DATA_BLOCK "DB149_KMI_FRA_Data"   // DB149
{ S7_Optimized_Access := 'FALSE' }
VERSION : 0.1
   VAR
      Signals_INT01 : Struct
         AP_ProgNr_Bit0 : Bool := FALSE;
         AP_ProgNr_Bit1 : Bool := FALSE;
         AP_ProgNr_Bit2 : Bool := FALSE;
         AP_ProgNr_Bit3 : Bool := FALSE;
         AP_ProgNr_Bit4 : Bool := FALSE;
         AP_ProgNr_Bit5 : Bool := FALSE;
         AP_ProgNr_Bit6 : Bool := FALSE;
         AP_ProgNr_Bit7 : Bool := FALSE;
         AP_OK : Bool := FALSE;
         AP_Strobe : Bool := FALSE;
         AP_Strobe_Inv : Bool := FALSE;
         AP_Shot : Bool := FALSE;
         AP_CP_forward : Bool := FALSE;
         AP_Filling : Bool := FALSE;
         AP_Res_0_6 : Bool := FALSE;
         AP_Res_0_7_1 : Bool := FALSE;
         PU_OK : Bool := FALSE;
         PU_Strobe_Quitt : Bool := FALSE;
         PU_Cycle_activ : Bool := FALSE;
         PU_Ready_for_shot : Bool := FALSE;
         PU_Shot_activ : Bool := FALSE;
         PU_Shot_End : Bool := FALSE;
         PU_Service_mode : Bool := TRUE;
         PU_CP_forward : Bool := FALSE;
         PU_Res_1_0 : Bool := FALSE;
         PU_Res_1_1 : Bool := FALSE;
         PU_Res_1_2 : Bool := FALSE;
         PU_Res_1_3 : Bool := FALSE;
         PU_Res_1_4 : Bool := FALSE;
         PU_Res_1_5 : Bool := FALSE;
         PU_Res_1_6 : Bool := FALSE;
         PU_Res_1_7 : Bool := FALSE;
         AP_Res_0_7 : Bool := FALSE;
      END_STRUCT;
      Measured_values_to_INT01 : Struct
         MH_Number : Byte := 16#01;
         Shot_Weight : Int := 16#1D40;
         Shot_Time : DInt := 16#0000_018D;
         Temperature_Poly : Int := 16#0794;
         Temperature_Iso : Int := 16#076C;
         Temperature_C3 : Int := 16#0000;
         Temperature_C4 : Int := 16#0000;
         Mix_Rate_Poly : Int := 16#2710;
         Mix_Rate_Iso : Int := 16#2F12;
         Mix_Rate_C3 : Int := 16#0000;
         Mix_Rate_C4 : Int := 16#0000;
         Pressure_Poly : Int := 16#466E;
         Pressure_Iso : Int := 16#44DE;
         Pressure_C3 : Int := 16#0000;
         Pressure_C4 : Int := 16#0000;
         Alarm_flow_K1 : Bool := FALSE;
         Alarm_flow_K2 : Bool := FALSE;
         Alarm_flow_K3 : Bool := FALSE;
         Alarm_flow_K4 : Bool := FALSE;
         Alarm_press_K1 : Bool := FALSE;
         Alarm_press_K2 : Bool := FALSE;
         Alarm_press_K3 : Bool := FALSE;
         Alarm_press_K4 : Bool := FALSE;
         Alarm_temp_K1 : Bool := FALSE;
         Alarm_temp_K2 : Bool := FALSE;
         Alarm_temp_K3 : Bool := FALSE;
         Alarm_temp_K4 : Bool := FALSE;
         Alarm_spare1 : Bool := FALSE;
         Alarm_spare2 : Bool := FALSE;
         Alarm_shottime : Bool := FALSE;
         Strobe_ProcessData : Bool := FALSE;
         Spare1 : Word := 16#0000;
         Spare2 : Word := 16#0000;
         Spare3 : Word := 16#0000;
         Spare4 : Word := 16#0000;
      END_STRUCT;
      Signals_INT02 : Struct
         AP_ProgNr_Bit0 : Bool := FALSE;
         AP_ProgNr_Bit1 : Bool := FALSE;
         AP_ProgNr_Bit2 : Bool := FALSE;
         AP_ProgNr_Bit3 : Bool := FALSE;
         AP_ProgNr_Bit4 : Bool := FALSE;
         AP_ProgNr_Bit5 : Bool := FALSE;
         AP_ProgNr_Bit6 : Bool := FALSE;
         AP_ProgNr_Bit7 : Bool := FALSE;
         AP_OK : Bool := FALSE;
         AP_Strobe : Bool := FALSE;
         AP_Strobe_Inv : Bool := FALSE;
         AP_Shot : Bool := FALSE;
         AP_CP_forward : Bool := FALSE;
         AP_Filling : Bool := FALSE;
         AP_Res_0_6 : Bool := FALSE;
         AP_Res_0_7_1 : Bool := FALSE;
         PU_OK : Bool := FALSE;
         PU_Strobe_Quitt : Bool := FALSE;
         PU_Cycle_activ : Bool := FALSE;
         PU_Ready_for_shot : Bool := FALSE;
         PU_Shot_activ : Bool := FALSE;
         PU_Shot_End : Bool := FALSE;
         PU_Service_mode : Bool := TRUE;
         PU_CP_forward : Bool := FALSE;
         PU_Res_1_0 : Bool := FALSE;
         PU_Res_1_1 : Bool := FALSE;
         PU_Res_1_2 : Bool := FALSE;
         PU_Res_1_3 : Bool := FALSE;
         PU_Res_1_4 : Bool := FALSE;
         PU_Res_1_5 : Bool := FALSE;
         PU_Res_1_6 : Bool := FALSE;
         PU_Res_1_7 : Bool := FALSE;
         AP_Res_0_7 : Bool := FALSE;
      END_STRUCT;
      Measured_values_to_INT02 : Struct
         MH_Number : Byte := 16#00;
         Shot_Weight : Int := 16#0000;
         Shot_Time : DInt := 16#0000_0000;
         Temperature_Poly : Int := 16#0000;
         Temperature_Iso : Int := 16#0000;
         Temperature_C3 : Int := 16#0000;
         Temperature_C4 : Int := 16#0000;
         Mix_Rate_Poly : Int := 16#0000;
         Mix_Rate_Iso : Int := 16#0000;
         Mix_Rate_C3 : Int := 16#0000;
         Mix_Rate_C4 : Int := 16#0000;
         Pressure_Poly : Int := 16#0000;
         Pressure_Iso : Int := 16#0000;
         Pressure_C3 : Int := 16#0000;
         Pressure_C4 : Int := 16#0000;
         Alarm_flow_K1 : Bool := FALSE;
         Alarm_flow_K2 : Bool := FALSE;
         Alarm_flow_K3 : Bool := FALSE;
         Alarm_flow_K4 : Bool := FALSE;
         Alarm_press_K1 : Bool := FALSE;
         Alarm_press_K2 : Bool := FALSE;
         Alarm_press_K3 : Bool := FALSE;
         Alarm_press_K4 : Bool := FALSE;
         Alarm_temp_K1 : Bool := FALSE;
         Alarm_temp_K2 : Bool := FALSE;
         Alarm_temp_K3 : Bool := FALSE;
         Alarm_temp_K4 : Bool := FALSE;
         Alarm_spare1 : Bool := FALSE;
         Alarm_spare2 : Bool := FALSE;
         Alarm_shottime : Bool := FALSE;
         Strobe_ProcessData : Bool := FALSE;
         Spare1 : Word := 16#0000;
         Spare2 : Word := 16#0000;
         Spare3 : Word := 16#0000;
         Spare4 : Word := 16#0000;
      END_STRUCT;
      Signals_INT03 : Struct
         AP_ProgNr_Bit0 : Bool := FALSE;
         AP_ProgNr_Bit1 : Bool := FALSE;
         AP_ProgNr_Bit2 : Bool := FALSE;
         AP_ProgNr_Bit3 : Bool := FALSE;
         AP_ProgNr_Bit4 : Bool := FALSE;
         AP_ProgNr_Bit5 : Bool := FALSE;
         AP_ProgNr_Bit6 : Bool := FALSE;
         AP_ProgNr_Bit7 : Bool := FALSE;
         AP_OK : Bool := FALSE;
         AP_Strobe : Bool := FALSE;
         AP_Strobe_Inv : Bool := FALSE;
         AP_Shot : Bool := FALSE;
         AP_CP_forward : Bool := FALSE;
         AP_Filling : Bool := FALSE;
         AP_Res_0_6 : Bool := FALSE;
         AP_Res_0_7_1 : Bool := FALSE;
         PU_OK : Bool := FALSE;
         PU_Strobe_Quitt : Bool := FALSE;
         PU_Cycle_activ : Bool := FALSE;
         PU_Ready_for_shot : Bool := FALSE;
         PU_Shot_activ : Bool := FALSE;
         PU_Shot_End : Bool := FALSE;
         PU_Service_mode : Bool := FALSE;
         PU_CP_forward : Bool := FALSE;
         PU_Res_1_0 : Bool := FALSE;
         PU_Res_1_1 : Bool := FALSE;
         PU_Res_1_2 : Bool := FALSE;
         PU_Res_1_3 : Bool := FALSE;
         PU_Res_1_4 : Bool := FALSE;
         PU_Res_1_5 : Bool := FALSE;
         PU_Res_1_6 : Bool := FALSE;
         PU_Res_1_7 : Bool := FALSE;
         AP_Res_0_7 : Bool := FALSE;
      END_STRUCT;
      Measured_values_to_INT03 : Struct
         MH_Number : Byte := 16#00;
         Shot_Weight : Int := 16#0000;
         Shot_Time : DInt := 16#0000_0000;
         Temperature_Poly : Int := 16#0000;
         Temperature_Iso : Int := 16#0000;
         Temperature_C3 : Int := 16#0000;
         Temperature_C4 : Int := 16#0000;
         Mix_Rate_Poly : Int := 16#0000;
         Mix_Rate_Iso : Int := 16#0000;
         Mix_Rate_C3 : Int := 16#0000;
         Mix_Rate_C4 : Int := 16#0000;
         Pressure_Poly : Int := 16#0000;
         Pressure_Iso : Int := 16#0000;
         Pressure_C3 : Int := 16#0000;
         Pressure_C4 : Int := 16#0000;
         Alarm_flow_K1 : Bool := FALSE;
         Alarm_flow_K2 : Bool := FALSE;
         Alarm_flow_K3 : Bool := FALSE;
         Alarm_flow_K4 : Bool := FALSE;
         Alarm_press_K1 : Bool := FALSE;
         Alarm_press_K2 : Bool := FALSE;
         Alarm_press_K3 : Bool := FALSE;
         Alarm_press_K4 : Bool := FALSE;
         Alarm_temp_K1 : Bool := FALSE;
         Alarm_temp_K2 : Bool := FALSE;
         Alarm_temp_K3 : Bool := FALSE;
         Alarm_temp_K4 : Bool := FALSE;
         Alarm_spare1 : Bool := FALSE;
         Alarm_spare2 : Bool := FALSE;
         Alarm_shottime : Bool := FALSE;
         Strobe_ProcessData : Bool := FALSE;
         Spare1 : Word := 16#0000;
         Spare2 : Word := 16#0000;
         Spare3 : Word := 16#0000;
         Spare4 : Word := 16#0000;
      END_STRUCT;
   END_VAR
BEGIN
END_DATA_BLOCK

DATA_BLOCK "DB_Zaehler_Anzeige"   // DB211
{ S7_Optimized_Access := 'FALSE' }
AUTHOR : AVP
NAME : MP270
VERSION : 0.1
   VAR
      ReadWriteDeviceNo : Int := 1;
      CopyDeviceNO : Int := 0;
      Read : Bool := FALSE;
      Write : Bool := FALSE;
      Copy : Bool := FALSE;
      Schichtwechsel : Bool := FALSE;
      ViewPreShift : Bool := FALSE;
      Gesamt : "Counter";
      "Counter" : Array[1..10] of "Counter";
      MH_Counter_ActualShift : Array[1..16] of Real;
      MH_Counter_PreShift : Array[1..16] of Real;
      MH_Counter_Reset : Array[1..16] of Real;
      MH_Counter_NonReset : Array[1..16] of Real;
   END_VAR
BEGIN
   Gesamt.Anzahl := 0;
   Gesamt.Verbrauch_K1 := 0.0;
   Gesamt.Verbrauch_K2 := 0.0;
   Gesamt.Verbrauch_K3 := 0.0;
   Gesamt.Verbrauch_K4 := 0.0;
   Gesamt.Verbrauch_K5 := 0.0;
   Gesamt.Verbrauch_K6 := 0.0;
   Gesamt.Verbrauch_K7 := 0.0;
   Gesamt.Verbrauch_K8 := 0.0;
   "Counter"[1].Anzahl := 0;
   "Counter"[1].Verbrauch_K1 := 0.0;
   "Counter"[1].Verbrauch_K2 := 0.0;
   "Counter"[1].Verbrauch_K3 := 0.0;
   "Counter"[1].Verbrauch_K4 := 0.0;
   "Counter"[1].Verbrauch_K5 := 0.0;
   "Counter"[1].Verbrauch_K6 := 0.0;
   "Counter"[1].Verbrauch_K7 := 0.0;
   "Counter"[1].Verbrauch_K8 := 0.0;
   "Counter"[2].Anzahl := 0;
   "Counter"[2].Verbrauch_K1 := 0.0;
   "Counter"[2].Verbrauch_K2 := 0.0;
   "Counter"[2].Verbrauch_K3 := 0.0;
   "Counter"[2].Verbrauch_K4 := 0.0;
   "Counter"[2].Verbrauch_K5 := 0.0;
   "Counter"[2].Verbrauch_K6 := 0.0;
   "Counter"[2].Verbrauch_K7 := 0.0;
   "Counter"[2].Verbrauch_K8 := 0.0;
   "Counter"[3].Anzahl := 0;
   "Counter"[3].Verbrauch_K1 := 0.0;
   "Counter"[3].Verbrauch_K2 := 0.0;
   "Counter"[3].Verbrauch_K3 := 0.0;
   "Counter"[3].Verbrauch_K4 := 0.0;
   "Counter"[3].Verbrauch_K5 := 0.0;
   "Counter"[3].Verbrauch_K6 := 0.0;
   "Counter"[3].Verbrauch_K7 := 0.0;
   "Counter"[3].Verbrauch_K8 := 0.0;
   "Counter"[4].Anzahl := 0;
   "Counter"[4].Verbrauch_K1 := 0.0;
   "Counter"[4].Verbrauch_K2 := 0.0;
   "Counter"[4].Verbrauch_K3 := 0.0;
   "Counter"[4].Verbrauch_K4 := 0.0;
   "Counter"[4].Verbrauch_K5 := 0.0;
   "Counter"[4].Verbrauch_K6 := 0.0;
   "Counter"[4].Verbrauch_K7 := 0.0;
   "Counter"[4].Verbrauch_K8 := 0.0;
   "Counter"[5].Anzahl := 0;
   "Counter"[5].Verbrauch_K1 := 0.0;
   "Counter"[5].Verbrauch_K2 := 0.0;
   "Counter"[5].Verbrauch_K3 := 0.0;
   "Counter"[5].Verbrauch_K4 := 0.0;
   "Counter"[5].Verbrauch_K5 := 0.0;
   "Counter"[5].Verbrauch_K6 := 0.0;
   "Counter"[5].Verbrauch_K7 := 0.0;
   "Counter"[5].Verbrauch_K8 := 0.0;
   "Counter"[6].Anzahl := 0;
   "Counter"[6].Verbrauch_K1 := 0.0;
   "Counter"[6].Verbrauch_K2 := 0.0;
   "Counter"[6].Verbrauch_K3 := 0.0;
   "Counter"[6].Verbrauch_K4 := 0.0;
   "Counter"[6].Verbrauch_K5 := 0.0;
   "Counter"[6].Verbrauch_K6 := 0.0;
   "Counter"[6].Verbrauch_K7 := 0.0;
   "Counter"[6].Verbrauch_K8 := 0.0;
   "Counter"[7].Anzahl := 0;
   "Counter"[7].Verbrauch_K1 := 0.0;
   "Counter"[7].Verbrauch_K2 := 0.0;
   "Counter"[7].Verbrauch_K3 := 0.0;
   "Counter"[7].Verbrauch_K4 := 0.0;
   "Counter"[7].Verbrauch_K5 := 0.0;
   "Counter"[7].Verbrauch_K6 := 0.0;
   "Counter"[7].Verbrauch_K7 := 0.0;
   "Counter"[7].Verbrauch_K8 := 0.0;
   "Counter"[8].Anzahl := 0;
   "Counter"[8].Verbrauch_K1 := 0.0;
   "Counter"[8].Verbrauch_K2 := 0.0;
   "Counter"[8].Verbrauch_K3 := 0.0;
   "Counter"[8].Verbrauch_K4 := 0.0;
   "Counter"[8].Verbrauch_K5 := 0.0;
   "Counter"[8].Verbrauch_K6 := 0.0;
   "Counter"[8].Verbrauch_K7 := 0.0;
   "Counter"[8].Verbrauch_K8 := 0.0;
   "Counter"[9].Anzahl := 0;
   "Counter"[9].Verbrauch_K1 := 0.0;
   "Counter"[9].Verbrauch_K2 := 0.0;
   "Counter"[9].Verbrauch_K3 := 0.0;
   "Counter"[9].Verbrauch_K4 := 0.0;
   "Counter"[9].Verbrauch_K5 := 0.0;
   "Counter"[9].Verbrauch_K6 := 0.0;
   "Counter"[9].Verbrauch_K7 := 0.0;
   "Counter"[9].Verbrauch_K8 := 0.0;
   "Counter"[10].Anzahl := 0;
   "Counter"[10].Verbrauch_K1 := 0.0;
   "Counter"[10].Verbrauch_K2 := 0.0;
   "Counter"[10].Verbrauch_K3 := 0.0;
   "Counter"[10].Verbrauch_K4 := 0.0;
   "Counter"[10].Verbrauch_K5 := 0.0;
   "Counter"[10].Verbrauch_K6 := 0.0;
   "Counter"[10].Verbrauch_K7 := 0.0;
   "Counter"[10].Verbrauch_K8 := 0.0;
   MH_Counter_ActualShift[1] := 0.0;
   MH_Counter_ActualShift[2] := 0.0;
   MH_Counter_ActualShift[3] := 0.0;
   MH_Counter_ActualShift[4] := 0.0;
   MH_Counter_ActualShift[5] := 0.0;
   MH_Counter_ActualShift[6] := 0.0;
   MH_Counter_ActualShift[7] := 0.0;
   MH_Counter_ActualShift[8] := 0.0;
   MH_Counter_ActualShift[9] := 0.0;
   MH_Counter_ActualShift[10] := 0.0;
   MH_Counter_ActualShift[11] := 0.0;
   MH_Counter_ActualShift[12] := 0.0;
   MH_Counter_ActualShift[13] := 0.0;
   MH_Counter_ActualShift[14] := 0.0;
   MH_Counter_ActualShift[15] := 0.0;
   MH_Counter_ActualShift[16] := 0.0;
   MH_Counter_PreShift[1] := 0.0;
   MH_Counter_PreShift[2] := 0.0;
   MH_Counter_PreShift[3] := 0.0;
   MH_Counter_PreShift[4] := 0.0;
   MH_Counter_PreShift[5] := 0.0;
   MH_Counter_PreShift[6] := 0.0;
   MH_Counter_PreShift[7] := 0.0;
   MH_Counter_PreShift[8] := 0.0;
   MH_Counter_PreShift[9] := 0.0;
   MH_Counter_PreShift[10] := 0.0;
   MH_Counter_PreShift[11] := 0.0;
   MH_Counter_PreShift[12] := 0.0;
   MH_Counter_PreShift[13] := 0.0;
   MH_Counter_PreShift[14] := 0.0;
   MH_Counter_PreShift[15] := 0.0;
   MH_Counter_PreShift[16] := 0.0;
   MH_Counter_Reset[1] := 0.0;
   MH_Counter_Reset[2] := 0.0;
   MH_Counter_Reset[3] := 0.0;
   MH_Counter_Reset[4] := 0.0;
   MH_Counter_Reset[5] := 0.0;
   MH_Counter_Reset[6] := 0.0;
   MH_Counter_Reset[7] := 0.0;
   MH_Counter_Reset[8] := 0.0;
   MH_Counter_Reset[9] := 0.0;
   MH_Counter_Reset[10] := 0.0;
   MH_Counter_Reset[11] := 0.0;
   MH_Counter_Reset[12] := 0.0;
   MH_Counter_Reset[13] := 0.0;
   MH_Counter_Reset[14] := 0.0;
   MH_Counter_Reset[15] := 0.0;
   MH_Counter_Reset[16] := 0.0;
   MH_Counter_NonReset[1] := 0.0;
   MH_Counter_NonReset[2] := 0.0;
   MH_Counter_NonReset[3] := 0.0;
   MH_Counter_NonReset[4] := 0.0;
   MH_Counter_NonReset[5] := 0.0;
   MH_Counter_NonReset[6] := 0.0;
   MH_Counter_NonReset[7] := 0.0;
   MH_Counter_NonReset[8] := 0.0;
   MH_Counter_NonReset[9] := 0.0;
   MH_Counter_NonReset[10] := 0.0;
   MH_Counter_NonReset[11] := 0.0;
   MH_Counter_NonReset[12] := 0.0;
   MH_Counter_NonReset[13] := 0.0;
   MH_Counter_NonReset[14] := 0.0;
   MH_Counter_NonReset[15] := 0.0;
   MH_Counter_NonReset[16] := 0.0;
END_DATA_BLOCK

DATA_BLOCK "DB_Zaehler_Schicht_aktuell"   // DB212
{ S7_Optimized_Access := 'FALSE' }
AUTHOR : AVP
NAME : MP270
VERSION : 0.1
   VAR
      Gesamt : "Counter";
      "Counter" : Array[1..120] of "Counter";
      MH_Counter : Array[1..16] of Real;
   END_VAR
BEGIN
   Gesamt.Anzahl := 0;
   Gesamt.Verbrauch_K1 := 0.0;
   Gesamt.Verbrauch_K2 := 0.0;
   Gesamt.Verbrauch_K3 := 0.0;
   Gesamt.Verbrauch_K4 := 0.0;
   Gesamt.Verbrauch_K5 := 0.0;
   Gesamt.Verbrauch_K6 := 0.0;
   Gesamt.Verbrauch_K7 := 0.0;
   Gesamt.Verbrauch_K8 := 0.0;
   "Counter"[1].Anzahl := 0;
   "Counter"[1].Verbrauch_K1 := 0.0;
   "Counter"[1].Verbrauch_K2 := 0.0;
   "Counter"[1].Verbrauch_K3 := 0.0;
   "Counter"[1].Verbrauch_K4 := 0.0;
   "Counter"[1].Verbrauch_K5 := 0.0;
   "Counter"[1].Verbrauch_K6 := 0.0;
   "Counter"[1].Verbrauch_K7 := 0.0;
   "Counter"[1].Verbrauch_K8 := 0.0;
   "Counter"[2].Anzahl := 0;
   "Counter"[2].Verbrauch_K1 := 0.0;
   "Counter"[2].Verbrauch_K2 := 0.0;
   "Counter"[2].Verbrauch_K3 := 0.0;
   "Counter"[2].Verbrauch_K4 := 0.0;
   "Counter"[2].Verbrauch_K5 := 0.0;
   "Counter"[2].Verbrauch_K6 := 0.0;
   "Counter"[2].Verbrauch_K7 := 0.0;
   "Counter"[2].Verbrauch_K8 := 0.0;
   "Counter"[3].Anzahl := 0;
   "Counter"[3].Verbrauch_K1 := 0.0;
   "Counter"[3].Verbrauch_K2 := 0.0;
   "Counter"[3].Verbrauch_K3 := 0.0;
   "Counter"[3].Verbrauch_K4 := 0.0;
   "Counter"[3].Verbrauch_K5 := 0.0;
   "Counter"[3].Verbrauch_K6 := 0.0;
   "Counter"[3].Verbrauch_K7 := 0.0;
   "Counter"[3].Verbrauch_K8 := 0.0;
   "Counter"[4].Anzahl := 0;
   "Counter"[4].Verbrauch_K1 := 0.0;
   "Counter"[4].Verbrauch_K2 := 0.0;
   "Counter"[4].Verbrauch_K3 := 0.0;
   "Counter"[4].Verbrauch_K4 := 0.0;
   "Counter"[4].Verbrauch_K5 := 0.0;
   "Counter"[4].Verbrauch_K6 := 0.0;
   "Counter"[4].Verbrauch_K7 := 0.0;
   "Counter"[4].Verbrauch_K8 := 0.0;
   "Counter"[5].Anzahl := 0;
   "Counter"[5].Verbrauch_K1 := 0.0;
   "Counter"[5].Verbrauch_K2 := 0.0;
   "Counter"[5].Verbrauch_K3 := 0.0;
   "Counter"[5].Verbrauch_K4 := 0.0;
   "Counter"[5].Verbrauch_K5 := 0.0;
   "Counter"[5].Verbrauch_K6 := 0.0;
   "Counter"[5].Verbrauch_K7 := 0.0;
   "Counter"[5].Verbrauch_K8 := 0.0;
   "Counter"[6].Anzahl := 0;
   "Counter"[6].Verbrauch_K1 := 0.0;
   "Counter"[6].Verbrauch_K2 := 0.0;
   "Counter"[6].Verbrauch_K3 := 0.0;
   "Counter"[6].Verbrauch_K4 := 0.0;
   "Counter"[6].Verbrauch_K5 := 0.0;
   "Counter"[6].Verbrauch_K6 := 0.0;
   "Counter"[6].Verbrauch_K7 := 0.0;
   "Counter"[6].Verbrauch_K8 := 0.0;
   "Counter"[7].Anzahl := 0;
   "Counter"[7].Verbrauch_K1 := 0.0;
   "Counter"[7].Verbrauch_K2 := 0.0;
   "Counter"[7].Verbrauch_K3 := 0.0;
   "Counter"[7].Verbrauch_K4 := 0.0;
   "Counter"[7].Verbrauch_K5 := 0.0;
   "Counter"[7].Verbrauch_K6 := 0.0;
   "Counter"[7].Verbrauch_K7 := 0.0;
   "Counter"[7].Verbrauch_K8 := 0.0;
   "Counter"[8].Anzahl := 0;
   "Counter"[8].Verbrauch_K1 := 0.0;
   "Counter"[8].Verbrauch_K2 := 0.0;
   "Counter"[8].Verbrauch_K3 := 0.0;
   "Counter"[8].Verbrauch_K4 := 0.0;
   "Counter"[8].Verbrauch_K5 := 0.0;
   "Counter"[8].Verbrauch_K6 := 0.0;
   "Counter"[8].Verbrauch_K7 := 0.0;
   "Counter"[8].Verbrauch_K8 := 0.0;
   "Counter"[9].Anzahl := 0;
   "Counter"[9].Verbrauch_K1 := 0.0;
   "Counter"[9].Verbrauch_K2 := 0.0;
   "Counter"[9].Verbrauch_K3 := 0.0;
   "Counter"[9].Verbrauch_K4 := 0.0;
   "Counter"[9].Verbrauch_K5 := 0.0;
   "Counter"[9].Verbrauch_K6 := 0.0;
   "Counter"[9].Verbrauch_K7 := 0.0;
   "Counter"[9].Verbrauch_K8 := 0.0;
   "Counter"[10].Anzahl := 0;
   "Counter"[10].Verbrauch_K1 := 0.0;
   "Counter"[10].Verbrauch_K2 := 0.0;
   "Counter"[10].Verbrauch_K3 := 0.0;
   "Counter"[10].Verbrauch_K4 := 0.0;
   "Counter"[10].Verbrauch_K5 := 0.0;
   "Counter"[10].Verbrauch_K6 := 0.0;
   "Counter"[10].Verbrauch_K7 := 0.0;
   "Counter"[10].Verbrauch_K8 := 0.0;
   "Counter"[11].Anzahl := 0;
   "Counter"[11].Verbrauch_K1 := 0.0;
   "Counter"[11].Verbrauch_K2 := 0.0;
   "Counter"[11].Verbrauch_K3 := 0.0;
   "Counter"[11].Verbrauch_K4 := 0.0;
   "Counter"[11].Verbrauch_K5 := 0.0;
   "Counter"[11].Verbrauch_K6 := 0.0;
   "Counter"[11].Verbrauch_K7 := 0.0;
   "Counter"[11].Verbrauch_K8 := 0.0;
   "Counter"[12].Anzahl := 0;
   "Counter"[12].Verbrauch_K1 := 0.0;
   "Counter"[12].Verbrauch_K2 := 0.0;
   "Counter"[12].Verbrauch_K3 := 0.0;
   "Counter"[12].Verbrauch_K4 := 0.0;
   "Counter"[12].Verbrauch_K5 := 0.0;
   "Counter"[12].Verbrauch_K6 := 0.0;
   "Counter"[12].Verbrauch_K7 := 0.0;
   "Counter"[12].Verbrauch_K8 := 0.0;
   "Counter"[13].Anzahl := 0;
   "Counter"[13].Verbrauch_K1 := 0.0;
   "Counter"[13].Verbrauch_K2 := 0.0;
   "Counter"[13].Verbrauch_K3 := 0.0;
   "Counter"[13].Verbrauch_K4 := 0.0;
   "Counter"[13].Verbrauch_K5 := 0.0;
   "Counter"[13].Verbrauch_K6 := 0.0;
   "Counter"[13].Verbrauch_K7 := 0.0;
   "Counter"[13].Verbrauch_K8 := 0.0;
   "Counter"[14].Anzahl := 0;
   "Counter"[14].Verbrauch_K1 := 0.0;
   "Counter"[14].Verbrauch_K2 := 0.0;
   "Counter"[14].Verbrauch_K3 := 0.0;
   "Counter"[14].Verbrauch_K4 := 0.0;
   "Counter"[14].Verbrauch_K5 := 0.0;
   "Counter"[14].Verbrauch_K6 := 0.0;
   "Counter"[14].Verbrauch_K7 := 0.0;
   "Counter"[14].Verbrauch_K8 := 0.0;
   "Counter"[15].Anzahl := 0;
   "Counter"[15].Verbrauch_K1 := 0.0;
   "Counter"[15].Verbrauch_K2 := 0.0;
   "Counter"[15].Verbrauch_K3 := 0.0;
   "Counter"[15].Verbrauch_K4 := 0.0;
   "Counter"[15].Verbrauch_K5 := 0.0;
   "Counter"[15].Verbrauch_K6 := 0.0;
   "Counter"[15].Verbrauch_K7 := 0.0;
   "Counter"[15].Verbrauch_K8 := 0.0;
   "Counter"[16].Anzahl := 0;
   "Counter"[16].Verbrauch_K1 := 0.0;
   "Counter"[16].Verbrauch_K2 := 0.0;
   "Counter"[16].Verbrauch_K3 := 0.0;
   "Counter"[16].Verbrauch_K4 := 0.0;
   "Counter"[16].Verbrauch_K5 := 0.0;
   "Counter"[16].Verbrauch_K6 := 0.0;
   "Counter"[16].Verbrauch_K7 := 0.0;
   "Counter"[16].Verbrauch_K8 := 0.0;
   "Counter"[17].Anzahl := 0;
   "Counter"[17].Verbrauch_K1 := 0.0;
   "Counter"[17].Verbrauch_K2 := 0.0;
   "Counter"[17].Verbrauch_K3 := 0.0;
   "Counter"[17].Verbrauch_K4 := 0.0;
   "Counter"[17].Verbrauch_K5 := 0.0;
   "Counter"[17].Verbrauch_K6 := 0.0;
   "Counter"[17].Verbrauch_K7 := 0.0;
   "Counter"[17].Verbrauch_K8 := 0.0;
   "Counter"[18].Anzahl := 0;
   "Counter"[18].Verbrauch_K1 := 0.0;
   "Counter"[18].Verbrauch_K2 := 0.0;
   "Counter"[18].Verbrauch_K3 := 0.0;
   "Counter"[18].Verbrauch_K4 := 0.0;
   "Counter"[18].Verbrauch_K5 := 0.0;
   "Counter"[18].Verbrauch_K6 := 0.0;
   "Counter"[18].Verbrauch_K7 := 0.0;
   "Counter"[18].Verbrauch_K8 := 0.0;
   "Counter"[19].Anzahl := 0;
   "Counter"[19].Verbrauch_K1 := 0.0;
   "Counter"[19].Verbrauch_K2 := 0.0;
   "Counter"[19].Verbrauch_K3 := 0.0;
   "Counter"[19].Verbrauch_K4 := 0.0;
   "Counter"[19].Verbrauch_K5 := 0.0;
   "Counter"[19].Verbrauch_K6 := 0.0;
   "Counter"[19].Verbrauch_K7 := 0.0;
   "Counter"[19].Verbrauch_K8 := 0.0;
   "Counter"[20].Anzahl := 0;
   "Counter"[20].Verbrauch_K1 := 0.0;
   "Counter"[20].Verbrauch_K2 := 0.0;
   "Counter"[20].Verbrauch_K3 := 0.0;
   "Counter"[20].Verbrauch_K4 := 0.0;
   "Counter"[20].Verbrauch_K5 := 0.0;
   "Counter"[20].Verbrauch_K6 := 0.0;
   "Counter"[20].Verbrauch_K7 := 0.0;
   "Counter"[20].Verbrauch_K8 := 0.0;
   "Counter"[21].Anzahl := 0;
   "Counter"[21].Verbrauch_K1 := 0.0;
   "Counter"[21].Verbrauch_K2 := 0.0;
   "Counter"[21].Verbrauch_K3 := 0.0;
   "Counter"[21].Verbrauch_K4 := 0.0;
   "Counter"[21].Verbrauch_K5 := 0.0;
   "Counter"[21].Verbrauch_K6 := 0.0;
   "Counter"[21].Verbrauch_K7 := 0.0;
   "Counter"[21].Verbrauch_K8 := 0.0;
   "Counter"[22].Anzahl := 0;
   "Counter"[22].Verbrauch_K1 := 0.0;
   // 905 more start values not shown
END_DATA_BLOCK

DATA_BLOCK "DB_Zaehler_Schicht_Vorherige"   // DB213
{ S7_Optimized_Access := 'FALSE' }
VERSION : 0.1
   VAR
      Gesamt : "Counter";
      "Counter" : Array[1..120] of "Counter";
      MH_Counter : Array[1..16] of Real;
   END_VAR
BEGIN
   Gesamt.Anzahl := 0;
   Gesamt.Verbrauch_K1 := 0.0;
   Gesamt.Verbrauch_K2 := 0.0;
   Gesamt.Verbrauch_K3 := 0.0;
   Gesamt.Verbrauch_K4 := 0.0;
   Gesamt.Verbrauch_K5 := 0.0;
   Gesamt.Verbrauch_K6 := 0.0;
   Gesamt.Verbrauch_K7 := 0.0;
   Gesamt.Verbrauch_K8 := 0.0;
   "Counter"[1].Anzahl := 0;
   "Counter"[1].Verbrauch_K1 := 0.0;
   "Counter"[1].Verbrauch_K2 := 0.0;
   "Counter"[1].Verbrauch_K3 := 0.0;
   "Counter"[1].Verbrauch_K4 := 0.0;
   "Counter"[1].Verbrauch_K5 := 0.0;
   "Counter"[1].Verbrauch_K6 := 0.0;
   "Counter"[1].Verbrauch_K7 := 0.0;
   "Counter"[1].Verbrauch_K8 := 0.0;
   "Counter"[2].Anzahl := 0;
   "Counter"[2].Verbrauch_K1 := 0.0;
   "Counter"[2].Verbrauch_K2 := 0.0;
   "Counter"[2].Verbrauch_K3 := 0.0;
   "Counter"[2].Verbrauch_K4 := 0.0;
   "Counter"[2].Verbrauch_K5 := 0.0;
   "Counter"[2].Verbrauch_K6 := 0.0;
   "Counter"[2].Verbrauch_K7 := 0.0;
   "Counter"[2].Verbrauch_K8 := 0.0;
   "Counter"[3].Anzahl := 0;
   "Counter"[3].Verbrauch_K1 := 0.0;
   "Counter"[3].Verbrauch_K2 := 0.0;
   "Counter"[3].Verbrauch_K3 := 0.0;
   "Counter"[3].Verbrauch_K4 := 0.0;
   "Counter"[3].Verbrauch_K5 := 0.0;
   "Counter"[3].Verbrauch_K6 := 0.0;
   "Counter"[3].Verbrauch_K7 := 0.0;
   "Counter"[3].Verbrauch_K8 := 0.0;
   "Counter"[4].Anzahl := 0;
   "Counter"[4].Verbrauch_K1 := 0.0;
   "Counter"[4].Verbrauch_K2 := 0.0;
   "Counter"[4].Verbrauch_K3 := 0.0;
   "Counter"[4].Verbrauch_K4 := 0.0;
   "Counter"[4].Verbrauch_K5 := 0.0;
   "Counter"[4].Verbrauch_K6 := 0.0;
   "Counter"[4].Verbrauch_K7 := 0.0;
   "Counter"[4].Verbrauch_K8 := 0.0;
   "Counter"[5].Anzahl := 0;
   "Counter"[5].Verbrauch_K1 := 0.0;
   "Counter"[5].Verbrauch_K2 := 0.0;
   "Counter"[5].Verbrauch_K3 := 0.0;
   "Counter"[5].Verbrauch_K4 := 0.0;
   "Counter"[5].Verbrauch_K5 := 0.0;
   "Counter"[5].Verbrauch_K6 := 0.0;
   "Counter"[5].Verbrauch_K7 := 0.0;
   "Counter"[5].Verbrauch_K8 := 0.0;
   "Counter"[6].Anzahl := 0;
   "Counter"[6].Verbrauch_K1 := 0.0;
   "Counter"[6].Verbrauch_K2 := 0.0;
   "Counter"[6].Verbrauch_K3 := 0.0;
   "Counter"[6].Verbrauch_K4 := 0.0;
   "Counter"[6].Verbrauch_K5 := 0.0;
   "Counter"[6].Verbrauch_K6 := 0.0;
   "Counter"[6].Verbrauch_K7 := 0.0;
   "Counter"[6].Verbrauch_K8 := 0.0;
   "Counter"[7].Anzahl := 0;
   "Counter"[7].Verbrauch_K1 := 0.0;
   "Counter"[7].Verbrauch_K2 := 0.0;
   "Counter"[7].Verbrauch_K3 := 0.0;
   "Counter"[7].Verbrauch_K4 := 0.0;
   "Counter"[7].Verbrauch_K5 := 0.0;
   "Counter"[7].Verbrauch_K6 := 0.0;
   "Counter"[7].Verbrauch_K7 := 0.0;
   "Counter"[7].Verbrauch_K8 := 0.0;
   "Counter"[8].Anzahl := 0;
   "Counter"[8].Verbrauch_K1 := 0.0;
   "Counter"[8].Verbrauch_K2 := 0.0;
   "Counter"[8].Verbrauch_K3 := 0.0;
   "Counter"[8].Verbrauch_K4 := 0.0;
   "Counter"[8].Verbrauch_K5 := 0.0;
   "Counter"[8].Verbrauch_K6 := 0.0;
   "Counter"[8].Verbrauch_K7 := 0.0;
   "Counter"[8].Verbrauch_K8 := 0.0;
   "Counter"[9].Anzahl := 0;
   "Counter"[9].Verbrauch_K1 := 0.0;
   "Counter"[9].Verbrauch_K2 := 0.0;
   "Counter"[9].Verbrauch_K3 := 0.0;
   "Counter"[9].Verbrauch_K4 := 0.0;
   "Counter"[9].Verbrauch_K5 := 0.0;
   "Counter"[9].Verbrauch_K6 := 0.0;
   "Counter"[9].Verbrauch_K7 := 0.0;
   "Counter"[9].Verbrauch_K8 := 0.0;
   "Counter"[10].Anzahl := 0;
   "Counter"[10].Verbrauch_K1 := 0.0;
   "Counter"[10].Verbrauch_K2 := 0.0;
   "Counter"[10].Verbrauch_K3 := 0.0;
   "Counter"[10].Verbrauch_K4 := 0.0;
   "Counter"[10].Verbrauch_K5 := 0.0;
   "Counter"[10].Verbrauch_K6 := 0.0;
   "Counter"[10].Verbrauch_K7 := 0.0;
   "Counter"[10].Verbrauch_K8 := 0.0;
   "Counter"[11].Anzahl := 0;
   "Counter"[11].Verbrauch_K1 := 0.0;
   "Counter"[11].Verbrauch_K2 := 0.0;
   "Counter"[11].Verbrauch_K3 := 0.0;
   "Counter"[11].Verbrauch_K4 := 0.0;
   "Counter"[11].Verbrauch_K5 := 0.0;
   "Counter"[11].Verbrauch_K6 := 0.0;
   "Counter"[11].Verbrauch_K7 := 0.0;
   "Counter"[11].Verbrauch_K8 := 0.0;
   "Counter"[12].Anzahl := 0;
   "Counter"[12].Verbrauch_K1 := 0.0;
   "Counter"[12].Verbrauch_K2 := 0.0;
   "Counter"[12].Verbrauch_K3 := 0.0;
   "Counter"[12].Verbrauch_K4 := 0.0;
   "Counter"[12].Verbrauch_K5 := 0.0;
   "Counter"[12].Verbrauch_K6 := 0.0;
   "Counter"[12].Verbrauch_K7 := 0.0;
   "Counter"[12].Verbrauch_K8 := 0.0;
   "Counter"[13].Anzahl := 0;
   "Counter"[13].Verbrauch_K1 := 0.0;
   "Counter"[13].Verbrauch_K2 := 0.0;
   "Counter"[13].Verbrauch_K3 := 0.0;
   "Counter"[13].Verbrauch_K4 := 0.0;
   "Counter"[13].Verbrauch_K5 := 0.0;
   "Counter"[13].Verbrauch_K6 := 0.0;
   "Counter"[13].Verbrauch_K7 := 0.0;
   "Counter"[13].Verbrauch_K8 := 0.0;
   "Counter"[14].Anzahl := 0;
   "Counter"[14].Verbrauch_K1 := 0.0;
   "Counter"[14].Verbrauch_K2 := 0.0;
   "Counter"[14].Verbrauch_K3 := 0.0;
   "Counter"[14].Verbrauch_K4 := 0.0;
   "Counter"[14].Verbrauch_K5 := 0.0;
   "Counter"[14].Verbrauch_K6 := 0.0;
   "Counter"[14].Verbrauch_K7 := 0.0;
   "Counter"[14].Verbrauch_K8 := 0.0;
   "Counter"[15].Anzahl := 0;
   "Counter"[15].Verbrauch_K1 := 0.0;
   "Counter"[15].Verbrauch_K2 := 0.0;
   "Counter"[15].Verbrauch_K3 := 0.0;
   "Counter"[15].Verbrauch_K4 := 0.0;
   "Counter"[15].Verbrauch_K5 := 0.0;
   "Counter"[15].Verbrauch_K6 := 0.0;
   "Counter"[15].Verbrauch_K7 := 0.0;
   "Counter"[15].Verbrauch_K8 := 0.0;
   "Counter"[16].Anzahl := 0;
   "Counter"[16].Verbrauch_K1 := 0.0;
   "Counter"[16].Verbrauch_K2 := 0.0;
   "Counter"[16].Verbrauch_K3 := 0.0;
   "Counter"[16].Verbrauch_K4 := 0.0;
   "Counter"[16].Verbrauch_K5 := 0.0;
   "Counter"[16].Verbrauch_K6 := 0.0;
   "Counter"[16].Verbrauch_K7 := 0.0;
   "Counter"[16].Verbrauch_K8 := 0.0;
   "Counter"[17].Anzahl := 0;
   "Counter"[17].Verbrauch_K1 := 0.0;
   "Counter"[17].Verbrauch_K2 := 0.0;
   "Counter"[17].Verbrauch_K3 := 0.0;
   "Counter"[17].Verbrauch_K4 := 0.0;
   "Counter"[17].Verbrauch_K5 := 0.0;
   "Counter"[17].Verbrauch_K6 := 0.0;
   "Counter"[17].Verbrauch_K7 := 0.0;
   "Counter"[17].Verbrauch_K8 := 0.0;
   "Counter"[18].Anzahl := 0;
   "Counter"[18].Verbrauch_K1 := 0.0;
   "Counter"[18].Verbrauch_K2 := 0.0;
   "Counter"[18].Verbrauch_K3 := 0.0;
   "Counter"[18].Verbrauch_K4 := 0.0;
   "Counter"[18].Verbrauch_K5 := 0.0;
   "Counter"[18].Verbrauch_K6 := 0.0;
   "Counter"[18].Verbrauch_K7 := 0.0;
   "Counter"[18].Verbrauch_K8 := 0.0;
   "Counter"[19].Anzahl := 0;
   "Counter"[19].Verbrauch_K1 := 0.0;
   "Counter"[19].Verbrauch_K2 := 0.0;
   "Counter"[19].Verbrauch_K3 := 0.0;
   "Counter"[19].Verbrauch_K4 := 0.0;
   "Counter"[19].Verbrauch_K5 := 0.0;
   "Counter"[19].Verbrauch_K6 := 0.0;
   "Counter"[19].Verbrauch_K7 := 0.0;
   "Counter"[19].Verbrauch_K8 := 0.0;
   "Counter"[20].Anzahl := 0;
   "Counter"[20].Verbrauch_K1 := 0.0;
   "Counter"[20].Verbrauch_K2 := 0.0;
   "Counter"[20].Verbrauch_K3 := 0.0;
   "Counter"[20].Verbrauch_K4 := 0.0;
   "Counter"[20].Verbrauch_K5 := 0.0;
   "Counter"[20].Verbrauch_K6 := 0.0;
   "Counter"[20].Verbrauch_K7 := 0.0;
   "Counter"[20].Verbrauch_K8 := 0.0;
   "Counter"[21].Anzahl := 0;
   "Counter"[21].Verbrauch_K1 := 0.0;
   "Counter"[21].Verbrauch_K2 := 0.0;
   "Counter"[21].Verbrauch_K3 := 0.0;
   "Counter"[21].Verbrauch_K4 := 0.0;
   "Counter"[21].Verbrauch_K5 := 0.0;
   "Counter"[21].Verbrauch_K6 := 0.0;
   "Counter"[21].Verbrauch_K7 := 0.0;
   "Counter"[21].Verbrauch_K8 := 0.0;
   "Counter"[22].Anzahl := 0;
   "Counter"[22].Verbrauch_K1 := 0.0;
   // 905 more start values not shown
END_DATA_BLOCK

DATA_BLOCK "DB315_ShotadjustS"   // DB315
TITLE = Shot time correction for each partshot of a tool
{ S7_Optimized_Access := 'FALSE' }
VERSION : 0.1
   VAR
      Tool : Array[0..120] of "UDT315_ShotadjustS";   // Shot time correction for each partshot of a tool
   END_VAR
BEGIN
   Tool[0].PS1 := 0.0;
END_DATA_BLOCK

DATA_BLOCK "DB601_PV_Plunger"   // DB601
TITLE = Process values of metering plunger
{ S7_Optimized_Access := 'FALSE' }
AUTHOR : KT242
VERSION : 0.1
   VAR
      ReadWriteDeviceNo : Int;
      CopyDeviceNO : Int;
      Read : Bool;
      Write : Bool;
      Copy : Bool;
      Component : Array[0..12] of "UDT509_PV_Plunger";
   END_VAR
BEGIN
END_DATA_BLOCK

DATA_BLOCK "DB602_PV_Tank"   // DB602
TITLE = Process values of tanks
{ S7_Optimized_Access := 'FALSE' }
AUTHOR : KT242